   3815: 'Spare_Fault_3815', class No Acknowledgement, trigger "DB302_HMI_Faults_Carrier59_Faults_2" bit 6
   3816: 'Spare_Fault_3816', class No Acknowledgement, trigger "DB302_HMI_Faults_Carrier59_Faults_2" bit 7
   3817: 'Spare_Fault_3817', class No Acknowledgement, trigger "DB302_HMI_Faults_Carrier59_Faults_2" bit 8
   3818: 'Spare_Fault_3818', class No Acknowledgement, trigger "DB302_HMI_Faults_Carrier59_Faults_2" bit 9
   3819: 'Spare_Fault_3819', class No Acknowledgement, trigger "DB302_HMI_Faults_Carrier59_Faults_2" bit 10
   3820: 'Spare_Fault_3820', class No Acknowledgement, trigger "DB302_HMI_Faults_Carrier59_Faults_2" bit 11
   3821: 'Spare_Fault_3821', class No Acknowledgement, trigger "DB302_HMI_Faults_Carrier59_Faults_2" bit 12
   3822: 'Spare_Fault_3822', class No Acknowledgement, trigger "DB302_HMI_Faults_Carrier59_Faults_2" bit 13
   3823: 'Spare_Fault_3823', class No Acknowledgement, trigger "DB302_HMI_Faults_Carrier59_Faults_2" bit 14
   3824: 'Spare_Fault_3824', class No Acknowledgement, trigger "DB302_HMI_Faults_Carrier59_Faults_2" bit 15
   3825: 'Spare_Fault_3825', class No Acknowledgement, trigger "DB302_HMI_Faults_Carrier59_Faults_3" bit 0
   3826: 'Spare_Fault_3826', class No Acknowledgement, trigger "DB302_HMI_Faults_Carrier59_Faults_3" bit 1
   3827: 'Spare_Fault_3827', class No Acknowledgement, trigger "DB302_HMI_Faults_Carrier59_Faults_3" bit 2
   3828: 'Spare_Fault_3828', class No Acknowledgement, trigger "DB302_HMI_Faults_Carrier59_Faults_3" bit 3
   3829: 'Spare_Fault_3829', class No Acknowledgement, trigger "DB302_HMI_Faults_Carrier59_Faults_3" bit 4
   3830: 'Spare_Fault_3830', class No Acknowledgement, trigger "DB302_HMI_Faults_Carrier59_Faults_3" bit 5
   3831: 'Spare_Fault_3831', class No Acknowledgement, trigger "DB302_HMI_Faults_Carrier59_Faults_3" bit 6
   3832: 'Spare_Fault_3832', class No Acknowledgement, trigger "DB302_HMI_Faults_Carrier59_Faults_3" bit 7
   3833: 'Spare_Fault_3833', class No Acknowledgement, trigger "DB302_HMI_Faults_Carrier59_Faults_3" bit 8
   3834: 'Spare_Fault_3834', class No Acknowledgement, trigger "DB302_HMI_Faults_Carrier59_Faults_3" bit 9
   3835: 'Spare_Fault_3835', class No Acknowledgement, trigger "DB302_HMI_Faults_Carrier59_Faults_3" bit 10
   3836: 'Spare_Fault_3836', class No Acknowledgement, trigger "DB302_HMI_Faults_Carrier59_Faults_3" bit 11
   3837: 'Spare_Fault_3837', class No Acknowledgement, trigger "DB302_HMI_Faults_Carrier59_Faults_3" bit 12
   3838: 'Spare_Fault_3838', class No Acknowledgement, trigger "DB302_HMI_Faults_Carrier59_Faults_3" bit 13
   3839: 'Spare_Fault_3839', class No Acknowledgement, trigger "DB302_HMI_Faults_Carrier59_Faults_3" bit 14
   3840: 'Spare_Fault_3840', class No Acknowledgement, trigger "DB302_HMI_Faults_Carrier59_Faults_3" bit 15
   3841: 'Carrier 60 Disconnect Open Power Fault DI11.0', class No Acknowledgement, trigger "DB302_HMI_Faults_Carrier60_Faults_0" bit 0
   3842: 'Carrier 60 Drive Profinet Comm Fault', class No Acknowledgement, trigger "DB302_HMI_Faults_Carrier60_Faults_0" bit 1
   3843: 'Carrier 60 Production Stop Not Reset', class No Acknowledgement, trigger "DB302_HMI_Faults_Carrier60_Faults_0" bit 2
   3844: 'Carrier 60 CB02122 Tripped', class No Acknowledgement, trigger "DB302_HMI_Faults_Carrier60_Faults_0" bit 3
   3845: 'Carrier 60 CB02123 Tripped', class No Acknowledgement, trigger "DB302_HMI_Faults_Carrier60_Faults_0" bit 4
   3846: 'Carrier 60 AUX1 CB Tripped', class No Acknowledgement, trigger "DB302_HMI_Faults_Carrier60_Faults_0" bit 5
   3847: 'Carrier 60 AUX2 CB Tripped', class No Acknowledgement, trigger "DB302_HMI_Faults_Carrier60_Faults_0" bit 6
   3848: 'Carrier 60 PLC Not Communicating', class No Acknowledgement, trigger "DB302_HMI_Faults_Carrier60_Faults_0" bit 7
   3849: 'Carrier 60 Safe Input Card Fault', class No Acknowledgement, trigger "DB302_HMI_Faults_Carrier60_Faults_0" bit 8
   3850: 'Carrier 60 Safe Output Card Fault', class No Acknowledgement, trigger "DB302_HMI_Faults_Carrier60_Faults_0" bit 9
   3851: 'Carrier 60 Standard Input Card Fault', class No Acknowledgement, trigger "DB302_HMI_Faults_Carrier60_Faults_0" bit 10
   3852: 'Carrier 60 Standard Output Card Fault', class No Acknowledgement, trigger "DB302_HMI_Faults_Carrier60_Faults_0" bit 11
   3853: 'Carrier 60 Encoder Position Fault', class No Acknowledgement, trigger "DB302_HMI_Faults_Carrier60_Faults_0" bit 12
   3854: 'Carrier 60 Encoder Internal Error', class No Acknowledgement, trigger "DB302_HMI_Faults_Carrier60_Faults_0" bit 13
   3855: 'Carrier 60 Encoder Comm Fault', class No Acknowledgement, trigger "DB302_HMI_Faults_Carrier60_Faults_0" bit 14
   3856: 'Carrier 60 HMI Comm Fault', class No Acknowledgement, trigger "DB302_HMI_Faults_Carrier60_Faults_0" bit 15
   3857: 'Carrier 60 Crash Detection Fault', class No Acknowledgement, trigger "DB302_HMI_Faults_Carrier60_Faults_1" bit 0
   3858: 'Carrier 60 Carrier Number Invalid', class No Acknowledgement, trigger "DB302_HMI_Faults_Carrier60_Faults_1" bit 1
   3859: 'Carrier 60 Drive: PROFINET configuration error', class No Acknowledgement, trigger "DB302_HMI_Faults_Carrier60_Faults_1" bit 2
   3860: 'Carrier 60 Drive: Error internal communications', class No Acknowledgement, trigger "DB302_HMI_Faults_Carrier60_Faults_1" bit 3
   3861: 'Carrier 60 Drive: Motor overtemperature', class No Acknowledgement, trigger "DB302_HMI_Faults_Carrier60_Faults_1" bit 4
   3862: 'Carrier 60 Drive: Motor overcurrent', class No Acknowledgement, trigger "DB302_HMI_Faults_Carrier60_Faults_1" bit 5
   3863: 'Carrier 60 Drive: Infeed or power unit not ready', class No Acknowledgement, trigger "DB302_HMI_Faults_Carrier60_Faults_1" bit 6
   3864: 'Carrier 60 Drive: Short-circuit/ground fault detected', class No Acknowledgement, trigger "DB302_HMI_Faults_Carrier60_Faults_1" bit 7
   3865: 'Carrier 60 Drive: PROFINET Setpoint timeout', class No Acknowledgement, trigger "DB302_HMI_Faults_Carrier60_Faults_1" bit 8
   3866: 'Carrier 60 Power unit: Overcurrent', class No Acknowledgement, trigger "DB302_HMI_Faults_Carrier60_Faults_1" bit 9
   3867: 'Carrier 60 Power unit: DC link voltage overvoltage', class No Acknowledgement, trigger "DB302_HMI_Faults_Carrier60_Faults_1" bit 10
   3868: 'Carrier 60 Power unit: DC link voltage undervoltage', class No Acknowledgement, trigger "DB302_HMI_Faults_Carrier60_Faults_1" bit 11
   3869: 'Carrier 60 Power unit: Line phase failure in main circuit', class No Acknowledgement, trigger "DB302_HMI_Faults_Carrier60_Faults_1" bit 12
   3870: 'Carrier 60 Power unit: Phase failure motor cable', class No Acknowledgement, trigger "DB302_HMI_Faults_Carrier60_Faults_1" bit 13
   3871: 'Carrier 60 Power unit: Ground fault', class No Acknowledgement, trigger "DB302_HMI_Faults_Carrier60_Faults_1" bit 14
   3872: 'Spare_Fault_3872', class No Acknowledgement, trigger "DB302_HMI_Faults_Carrier60_Faults_1" bit 15
   3873: 'Carrier 60 Motion Off Fault', class No Acknowledgement, trigger "DB302_HMI_Faults_Carrier60_Faults_2" bit 0
   3874: 'Carrier 60 Motion On Fault', class No Acknowledgement, trigger "DB302_HMI_Faults_Carrier60_Faults_2" bit 1
   3875: 'Carrier 60 Spacing Fault', class No Acknowledgement, trigger "DB302_HMI_Faults_Carrier60_Faults_2" bit 2
   3876: 'Carrier 60 Duplicate Carrier Number Fault', class No Acknowledgement, trigger "DB302_HMI_Faults_Carrier60_Faults_2" bit 3
   3877: 'Spare_Fault_3877', class No Acknowledgement, trigger "DB302_HMI_Faults_Carrier60_Faults_2" bit 4
   3878: 'Spare_Fault_3878', class No Acknowledgement, trigger "DB302_HMI_Faults_Carrier60_Faults_2" bit 5
   3879: 'Spare_Fault_3879', class No Acknowledgement, trigger "DB302_HMI_Faults_Carrier60_Faults_2" bit 6
   3880: 'Spare_Fault_3880', class No Acknowledgement, trigger "DB302_HMI_Faults_Carrier60_Faults_2" bit 7
   3881: 'Spare_Fault_3881', class No Acknowledgement, trigger "DB302_HMI_Faults_Carrier60_Faults_2" bit 8
   3882: 'Spare_Fault_3882', class No Acknowledgement, trigger "DB302_HMI_Faults_Carrier60_Faults_2" bit 9
   3883: 'Spare_Fault_3883', class No Acknowledgement, trigger "DB302_HMI_Faults_Carrier60_Faults_2" bit 10
   3884: 'Spare_Fault_3884', class No Acknowledgement, trigger "DB302_HMI_Faults_Carrier60_Faults_2" bit 11
   3885: 'Spare_Fault_3885', class No Acknowledgement, trigger "DB302_HMI_Faults_Carrier60_Faults_2" bit 12
   3886: 'Spare_Fault_3886', class No Acknowledgement, trigger "DB302_HMI_Faults_Carrier60_Faults_2" bit 13
   3887: 'Spare_Fault_3887', class No Acknowledgement, trigger "DB302_HMI_Faults_Carrier60_Faults_2" bit 14
   3888: 'Spare_Fault_3888', class No Acknowledgement, trigger "DB302_HMI_Faults_Carrier60_Faults_2" bit 15
   3889: 'Spare_Fault_3889', class No Acknowledgement, trigger "DB302_HMI_Faults_Carrier60_Faults_3" bit 0
   3890: 'Spare_Fault_3890', class No Acknowledgement, trigger "DB302_HMI_Faults_Carrier60_Faults_3" bit 1
   3891: 'Spare_Fault_3891', class No Acknowledgement, trigger "DB302_HMI_Faults_Carrier60_Faults_3" bit 2
   3892: 'Spare_Fault_3892', class No Acknowledgement, trigger "DB302_HMI_Faults_Carrier60_Faults_3" bit 3
   3893: 'Spare_Fault_3893', class No Acknowledgement, trigger "DB302_HMI_Faults_Carrier60_Faults_3" bit 4
   3894: 'Spare_Fault_3894', class No Acknowledgement, trigger "DB302_HMI_Faults_Carrier60_Faults_3" bit 5
   3895: 'Spare_Fault_3895', class No Acknowledgement, trigger "DB302_HMI_Faults_Carrier60_Faults_3" bit 6
   3896: 'Spare_Fault_3896', class No Acknowledgement, trigger "DB302_HMI_Faults_Carrier60_Faults_3" bit 7
   3897: 'Spare_Fault_3897', class No Acknowledgement, trigger "DB302_HMI_Faults_Carrier60_Faults_3" bit 8
   3898: 'Spare_Fault_3898', class No Acknowledgement, trigger "DB302_HMI_Faults_Carrier60_Faults_3" bit 9
   3899: 'Spare_Fault_3899', class No Acknowledgement, trigger "DB302_HMI_Faults_Carrier60_Faults_3" bit 10
   3900: 'Spare_Fault_3900', class No Acknowledgement, trigger "DB302_HMI_Faults_Carrier60_Faults_3" bit 11
   3901: 'Spare_Fault_3901', class No Acknowledgement, trigger "DB302_HMI_Faults_Carrier60_Faults_3" bit 12
   3902: 'Spare_Fault_3902', class No Acknowledgement, trigger "DB302_HMI_Faults_Carrier60_Faults_3" bit 13
   3903: 'Spare_Fault_3903', class No Acknowledgement, trigger "DB302_HMI_Faults_Carrier60_Faults_3" bit 14
   3904: 'Spare_Fault_3904', class No Acknowledgement, trigger "DB302_HMI_Faults_Carrier60_Faults_3" bit 15
   3905: 'Carrier 61 Disconnect Open Power Fault DI11.0', class No Acknowledgement, trigger "DB302_HMI_Faults_Carrier61_Faults_0" bit 0
   3906: 'Carrier 61 Drive Profinet Comm Fault', class No Acknowledgement, trigger "DB302_HMI_Faults_Carrier61_Faults_0" bit 1
   3907: 'Carrier 61 Production Stop Not Reset', class No Acknowledgement, trigger "DB302_HMI_Faults_Carrier61_Faults_0" bit 2
   3908: 'Carrier 61 CB02122 Tripped', class No Acknowledgement, trigger "DB302_HMI_Faults_Carrier61_Faults_0" bit 3
   3909: 'Carrier 61 CB02123 Tripped', class No Acknowledgement, trigger "DB302_HMI_Faults_Carrier61_Faults_0" bit 4
   3910: 'Carrier 61 AUX1 CB Tripped', class No Acknowledgement, trigger "DB302_HMI_Faults_Carrier61_Faults_0" bit 5
   3911: 'Carrier 61 AUX2 CB Tripped', class No Acknowledgement, trigger "DB302_HMI_Faults_Carrier61_Faults_0" bit 6
   3912: 'Carrier 61 PLC Not Communicating', class No Acknowledgement, trigger "DB302_HMI_Faults_Carrier61_Faults_0" bit 7
   3913: 'Carrier 61 Safe Input Card Fault', class No Acknowledgement, trigger "DB302_HMI_Faults_Carrier61_Faults_0" bit 8
   3914: 'Carrier 61 Safe Output Card Fault', class No Acknowledgement, trigger "DB302_HMI_Faults_Carrier61_Faults_0" bit 9
   3915: 'Carrier 61 Standard Input Card Fault', class No Acknowledgement, trigger "DB302_HMI_Faults_Carrier61_Faults_0" bit 10
   3916: 'Carrier 61 Standard Output Card Fault', class No Acknowledgement, trigger "DB302_HMI_Faults_Carrier61_Faults_0" bit 11
   3917: 'Carrier 61 Encoder Position Fault', class No Acknowledgement, trigger "DB302_HMI_Faults_Carrier61_Faults_0" bit 12
   3918: 'Carrier 61 Encoder Internal Error', class No Acknowledgement, trigger "DB302_HMI_Faults_Carrier61_Faults_0" bit 13
   3919: 'Carrier 61 Encoder Comm Fault', class No Acknowledgement, trigger "DB302_HMI_Faults_Carrier61_Faults_0" bit 14
   3920: 'Carrier 61 HMI Comm Fault', class No Acknowledgement, trigger "DB302_HMI_Faults_Carrier61_Faults_0" bit 15
   3921: 'Carrier 61 Crash Detection Fault', class No Acknowledgement, trigger "DB302_HMI_Faults_Carrier61_Faults_1" bit 0
   3922: 'Carrier 61 Carrier Number Invalid', class No Acknowledgement, trigger "DB302_HMI_Faults_Carrier61_Faults_1" bit 1
   3923: 'Carrier 61 Drive: PROFINET configuration error', class No Acknowledgement, trigger "DB302_HMI_Faults_Carrier61_Faults_1" bit 2
   3924: 'Carrier 61 Drive: Error internal communications', class No Acknowledgement, trigger "DB302_HMI_Faults_Carrier61_Faults_1" bit 3
   3925: 'Carrier 61 Drive: Motor overtemperature', class No Acknowledgement, trigger "DB302_HMI_Faults_Carrier61_Faults_1" bit 4
   3926: 'Carrier 61 Drive: Motor overcurrent', class No Acknowledgement, trigger "DB302_HMI_Faults_Carrier61_Faults_1" bit 5
   3927: 'Carrier 61 Drive: Infeed or power unit not ready', class No Acknowledgement, trigger "DB302_HMI_Faults_Carrier61_Faults_1" bit 6
   3928: 'Carrier 61 Drive: Short-circuit/ground fault detected', class No Acknowledgement, trigger "DB302_HMI_Faults_Carrier61_Faults_1" bit 7
   3929: 'Carrier 61 Drive: PROFINET Setpoint timeout', class No Acknowledgement, trigger "DB302_HMI_Faults_Carrier61_Faults_1" bit 8
   3930: 'Carrier 61 Power unit: Overcurrent', class No Acknowledgement, trigger "DB302_HMI_Faults_Carrier61_Faults_1" bit 9
   3931: 'Carrier 61 Power unit: DC link voltage overvoltage', class No Acknowledgement, trigger "DB302_HMI_Faults_Carrier61_Faults_1" bit 10
   3932: 'Carrier 61 Power unit: DC link voltage undervoltage', class No Acknowledgement, trigger "DB302_HMI_Faults_Carrier61_Faults_1" bit 11
   3933: 'Carrier 61 Power unit: Line phase failure in main circuit', class No Acknowledgement, trigger "DB302_HMI_Faults_Carrier61_Faults_1" bit 12
   3934: 'Carrier 61 Power unit: Phase failure motor cable', class No Acknowledgement, trigger "DB302_HMI_Faults_Carrier61_Faults_1" bit 13
   3935: 'Carrier 61 Power unit: Ground fault', class No Acknowledgement, trigger "DB302_HMI_Faults_Carrier61_Faults_1" bit 14
   3936: 'Spare_Fault_3936', class No Acknowledgement, trigger "DB302_HMI_Faults_Carrier61_Faults_1" bit 15
   3937: 'Carrier 61 Motion Off Fault', class No Acknowledgement, trigger "DB302_HMI_Faults_Carrier61_Faults_2" bit 0
   3938: 'Carrier 61 Motion On Fault', class No Acknowledgement, trigger "DB302_HMI_Faults_Carrier61_Faults_2" bit 1
   3939: 'Carrier 61 Spacing Fault', class No Acknowledgement, trigger "DB302_HMI_Faults_Carrier61_Faults_2" bit 2
   3940: 'Carrier 61 Duplicate Carrier Number Fault', class No Acknowledgement, trigger "DB302_HMI_Faults_Carrier61_Faults_2" bit 3
   3941: 'Spare_Fault_3941', class No Acknowledgement, trigger "DB302_HMI_Faults_Carrier61_Faults_2" bit 4
   3942: 'Spare_Fault_3942', class No Acknowledgement, trigger "DB302_HMI_Faults_Carrier61_Faults_2" bit 5
   3943: 'Spare_Fault_3943', class No Acknowledgement, trigger "DB302_HMI_Faults_Carrier61_Faults_2" bit 6
   3944: 'Spare_Fault_3944', class No Acknowledgement, trigger "DB302_HMI_Faults_Carrier61_Faults_2" bit 7
   3945: 'Spare_Fault_3945', class No Acknowledgement, trigger "DB302_HMI_Faults_Carrier61_Faults_2" bit 8
   3946: 'Spare_Fault_3946', class No Acknowledgement, trigger "DB302_HMI_Faults_Carrier61_Faults_2" bit 9
   3947: 'Spare_Fault_3947', class No Acknowledgement, trigger "DB302_HMI_Faults_Carrier61_Faults_2" bit 10
   3948: 'Spare_Fault_3948', class No Acknowledgement, trigger "DB302_HMI_Faults_Carrier61_Faults_2" bit 11
   3949: 'Spare_Fault_3949', class No Acknowledgement, trigger "DB302_HMI_Faults_Carrier61_Faults_2" bit 12
   3950: 'Spare_Fault_3950', class No Acknowledgement, trigger "DB302_HMI_Faults_Carrier61_Faults_2" bit 13
   3951: 'Spare_Fault_3951', class No Acknowledgement, trigger "DB302_HMI_Faults_Carrier61_Faults_2" bit 14
   3952: 'Spare_Fault_3952', class No Acknowledgement, trigger "DB302_HMI_Faults_Carrier61_Faults_2" bit 15
   3953: 'Spare_Fault_3953', class No Acknowledgement, trigger "DB302_HMI_Faults_Carrier61_Faults_3" bit 0
   3954: 'Spare_Fault_3954', class No Acknowledgement, trigger "DB302_HMI_Faults_Carrier61_Faults_3" bit 1
   3955: 'Spare_Fault_3955', class No Acknowledgement, trigger "DB302_HMI_Faults_Carrier61_Faults_3" bit 2
   3956: 'Spare_Fault_3956', class No Acknowledgement, trigger "DB302_HMI_Faults_Carrier61_Faults_3" bit 3
   3957: 'Spare_Fault_3957', class No Acknowledgement, trigger "DB302_HMI_Faults_Carrier61_Faults_3" bit 4
   3958: 'Spare_Fault_3958', class No Acknowledgement, trigger "DB302_HMI_Faults_Carrier61_Faults_3" bit 5
   3959: 'Spare_Fault_3959', class No Acknowledgement, trigger "DB302_HMI_Faults_Carrier61_Faults_3" bit 6
   3960: 'Spare_Fault_3960', class No Acknowledgement, trigger "DB302_HMI_Faults_Carrier61_Faults_3" bit 7
   3961: 'Spare_Fault_3961', class No Acknowledgement, trigger "DB302_HMI_Faults_Carrier61_Faults_3" bit 8
   3962: 'Spare_Fault_3962', class No Acknowledgement, trigger "DB302_HMI_Faults_Carrier61_Faults_3" bit 9
   3963: 'Spare_Fault_3963', class No Acknowledgement, trigger "DB302_HMI_Faults_Carrier61_Faults_3" bit 10
   3964: 'Spare_Fault_3964', class No Acknowledgement, trigger "DB302_HMI_Faults_Carrier61_Faults_3" bit 11
   3965: 'Spare_Fault_3965', class No Acknowledgement, trigger "DB302_HMI_Faults_Carrier61_Faults_3" bit 12
   3966: 'Spare_Fault_3966', class No Acknowledgement, trigger "DB302_HMI_Faults_Carrier61_Faults_3" bit 13
   3967: 'Spare_Fault_3967', class No Acknowledgement, trigger "DB302_HMI_Faults_Carrier61_Faults_3" bit 14
   3968: 'Spare_Fault_3968', class No Acknowledgement, trigger "DB302_HMI_Faults_Carrier61_Faults_3" bit 15
   3969: 'Carrier 62 Disconnect Open Power Fault DI11.0', class No Acknowledgement, trigger "DB302_HMI_Faults_Carrier62_Faults_0" bit 0
   3970: 'Carrier 62 Drive Profinet Comm Fault', class No Acknowledgement, trigger "DB302_HMI_Faults_Carrier62_Faults_0" bit 1
   3971: 'Carrier 62 Production Stop Not Reset', class No Acknowledgement, trigger "DB302_HMI_Faults_Carrier62_Faults_0" bit 2
   3972: 'Carrier 62 CB02122 Tripped', class No Acknowledgement, trigger "DB302_HMI_Faults_Carrier62_Faults_0" bit 3
   3973: 'Carrier 62 CB02123 Tripped', class No Acknowledgement, trigger "DB302_HMI_Faults_Carrier62_Faults_0" bit 4
   3974: 'Carrier 62 AUX1 CB Tripped', class No Acknowledgement, trigger "DB302_HMI_Faults_Carrier62_Faults_0" bit 5
   3975: 'Carrier 62 AUX2 CB Tripped', class No Acknowledgement, trigger "DB302_HMI_Faults_Carrier62_Faults_0" bit 6
   3976: 'Carrier 62 PLC Not Communicating', class No Acknowledgement, trigger "DB302_HMI_Faults_Carrier62_Faults_0" bit 7
   3977: 'Carrier 62 Safe Input Card Fault', class No Acknowledgement, trigger "DB302_HMI_Faults_Carrier62_Faults_0" bit 8
   3978: 'Carrier 62 Safe Output Card Fault', class No Acknowledgement, trigger "DB302_HMI_Faults_Carrier62_Faults_0" bit 9
   3979: 'Carrier 62 Standard Input Card Fault', class No Acknowledgement, trigger "DB302_HMI_Faults_Carrier62_Faults_0" bit 10
   3980: 'Carrier 62 Standard Output Card Fault', class No Acknowledgement, trigger "DB302_HMI_Faults_Carrier62_Faults_0" bit 11
   3981: 'Carrier 62 Encoder Position Fault', class No Acknowledgement, trigger "DB302_HMI_Faults_Carrier62_Faults_0" bit 12
   3982: 'Carrier 62 Encoder Internal Error', class No Acknowledgement, trigger "DB302_HMI_Faults_Carrier62_Faults_0" bit 13
   3983: 'Carrier 62 Encoder Comm Fault', class No Acknowledgement, trigger "DB302_HMI_Faults_Carrier62_Faults_0" bit 14
   3984: 'Carrier 62 HMI Comm Fault', class No Acknowledgement, trigger "DB302_HMI_Faults_Carrier62_Faults_0" bit 15
   3985: 'Carrier 62 Crash Detection Fault', class No Acknowledgement, trigger "DB302_HMI_Faults_Carrier62_Faults_1" bit 0
   3986: 'Carrier 62 Carrier Number Invalid', class No Acknowledgement, trigger "DB302_HMI_Faults_Carrier62_Faults_1" bit 1
   3987: 'Carrier 62 Drive: PROFINET configuration error', class No Acknowledgement, trigger "DB302_HMI_Faults_Carrier62_Faults_1" bit 2
   3988: 'Carrier 62 Drive: Error internal communications', class No Acknowledgement, trigger "DB302_HMI_Faults_Carrier62_Faults_1" bit 3
   3989: 'Carrier 62 Drive: Motor overtemperature', class No Acknowledgement, trigger "DB302_HMI_Faults_Carrier62_Faults_1" bit 4
   3990: 'Carrier 62 Drive: Motor overcurrent', class No Acknowledgement, trigger "DB302_HMI_Faults_Carrier62_Faults_1" bit 5
   3991: 'Carrier 62 Drive: Infeed or power unit not ready', class No Acknowledgement, trigger "DB302_HMI_Faults_Carrier62_Faults_1" bit 6
   3992: 'Carrier 62 Drive: Short-circuit/ground fault detected', class No Acknowledgement, trigger "DB302_HMI_Faults_Carrier62_Faults_1" bit 7
   3993: 'Carrier 62 Drive: PROFINET Setpoint timeout', class No Acknowledgement, trigger "DB302_HMI_Faults_Carrier62_Faults_1" bit 8
   3994: 'Carrier 62 Power unit: Overcurrent', class No Acknowledgement, trigger "DB302_HMI_Faults_Carrier62_Faults_1" bit 9
   3995: 'Carrier 62 Power unit: DC link voltage overvoltage', class No Acknowledgement, trigger "DB302_HMI_Faults_Carrier62_Faults_1" bit 10
   3996: 'Carrier 62 Power unit: DC link voltage undervoltage', class No Acknowledgement, trigger "DB302_HMI_Faults_Carrier62_Faults_1" bit 11
   3997: 'Carrier 62 Power unit: Line phase failure in main circuit', class No Acknowledgement, trigger "DB302_HMI_Faults_Carrier62_Faults_1" bit 12
   3998: 'Carrier 62 Power unit: Phase failure motor cable', class No Acknowledgement, trigger "DB302_HMI_Faults_Carrier62_Faults_1" bit 13
   3999: 'Carrier 62 Power unit: Ground fault', class No Acknowledgement, trigger "DB302_HMI_Faults_Carrier62_Faults_1" bit 14
   4000: 'Spare_Fault_4000', class No Acknowledgement, trigger "DB302_HMI_Faults_Carrier62_Faults_1" bit 15
   4001: 'Carrier 62 Motion Off Fault', class No Acknowledgement, trigger "DB302_HMI_Faults_Carrier62_Faults_2" bit 0
   4002: 'Carrier 62 Motion On Fault', class No Acknowledgement, trigger "DB302_HMI_Faults_Carrier62_Faults_2" bit 1
   4003: 'Carrier 62 Spacing Fault', class No Acknowledgement, trigger "DB302_HMI_Faults_Carrier62_Faults_2" bit 2
   4004: 'Carrier 62 Duplicate Carrier Number Fault', class No Acknowledgement, trigger "DB302_HMI_Faults_Carrier62_Faults_2" bit 3
   4005: 'Spare_Fault_4005', class No Acknowledgement, trigger "DB302_HMI_Faults_Carrier62_Faults_2" bit 4
   4006: 'Spare_Fault_4006', class No Acknowledgement, trigger "DB302_HMI_Faults_Carrier62_Faults_2" bit 5
   4007: 'Spare_Fault_4007', class No Acknowledgement, trigger "DB302_HMI_Faults_Carrier62_Faults_2" bit 6
   4008: 'Spare_Fault_4008', class No Acknowledgement, trigger "DB302_HMI_Faults_Carrier62_Faults_2" bit 7
   4009: 'Spare_Fault_4009', class No Acknowledgement, trigger "DB302_HMI_Faults_Carrier62_Faults_2" bit 8
   4010: 'Spare_Fault_4010', class No Acknowledgement, trigger "DB302_HMI_Faults_Carrier62_Faults_2" bit 9
   4011: 'Spare_Fault_4011', class No Acknowledgement, trigger "DB302_HMI_Faults_Carrier62_Faults_2" bit 10
   4012: 'Spare_Fault_4012', class No Acknowledgement, trigger "DB302_HMI_Faults_Carrier62_Faults_2" bit 11
   4013: 'Spare_Fault_4013', class No Acknowledgement, trigger "DB302_HMI_Faults_Carrier62_Faults_2" bit 12
   4014: 'Spare_Fault_4014', class No Acknowledgement, trigger "DB302_HMI_Faults_Carrier62_Faults_2" bit 13
   4015: 'Spare_Fault_4015', class No Acknowledgement, trigger "DB302_HMI_Faults_Carrier62_Faults_2" bit 14
   4016: 'Spare_Fault_4016', class No Acknowledgement, trigger "DB302_HMI_Faults_Carrier62_Faults_2" bit 15
   4017: 'Spare_Fault_4017', class No Acknowledgement, trigger "DB302_HMI_Faults_Carrier62_Faults_3" bit 0
   4018: 'Spare_Fault_4018', class No Acknowledgement, trigger "DB302_HMI_Faults_Carrier62_Faults_3" bit 1
   4019: 'Spare_Fault_4019', class No Acknowledgement, trigger "DB302_HMI_Faults_Carrier62_Faults_3" bit 2
   4020: 'Spare_Fault_4020', class No Acknowledgement, trigger "DB302_HMI_Faults_Carrier62_Faults_3" bit 3
   4021: 'Spare_Fault_4021', class No Acknowledgement, trigger "DB302_HMI_Faults_Carrier62_Faults_3" bit 4
   4022: 'Spare_Fault_4022', class No Acknowledgement, trigger "DB302_HMI_Faults_Carrier62_Faults_3" bit 5
   4023: 'Spare_Fault_4023', class No Acknowledgement, trigger "DB302_HMI_Faults_Carrier62_Faults_3" bit 6
   4024: 'Spare_Fault_4024', class No Acknowledgement, trigger "DB302_HMI_Faults_Carrier62_Faults_3" bit 7
   4025: 'Spare_Fault_4025', class No Acknowledgement, trigger "DB302_HMI_Faults_Carrier62_Faults_3" bit 8
   4026: 'Spare_Fault_4026', class No Acknowledgement, trigger "DB302_HMI_Faults_Carrier62_Faults_3" bit 9
   4027: 'Spare_Fault_4027', class No Acknowledgement, trigger "DB302_HMI_Faults_Carrier62_Faults_3" bit 10
   4028: 'Spare_Fault_4028', class No Acknowledgement, trigger "DB302_HMI_Faults_Carrier62_Faults_3" bit 11
   4029: 'Spare_Fault_4029', class No Acknowledgement, trigger "DB302_HMI_Faults_Carrier62_Faults_3" bit 12
   4030: 'Spare_Fault_4030', class No Acknowledgement, trigger "DB302_HMI_Faults_Carrier62_Faults_3" bit 13
   4031: 'Spare_Fault_4031', class No Acknowledgement, trigger "DB302_HMI_Faults_Carrier62_Faults_3" bit 14
   4032: 'Spare_Fault_4032', class No Acknowledgement, trigger "DB302_HMI_Faults_Carrier62_Faults_3" bit 15
   4033: 'Carrier 63 Disconnect Open Power Fault DI11.0', class No Acknowledgement, trigger "DB302_HMI_Faults_Carrier63_Faults_0" bit 0
   4034: 'Carrier 63 Drive Profinet Comm Fault', class No Acknowledgement, trigger "DB302_HMI_Faults_Carrier63_Faults_0" bit 1
   4035: 'Carrier 63 Production Stop Not Reset', class No Acknowledgement, trigger "DB302_HMI_Faults_Carrier63_Faults_0" bit 2
   4036: 'Carrier 63 CB02122 Tripped', class No Acknowledgement, trigger "DB302_HMI_Faults_Carrier63_Faults_0" bit 3
   4037: 'Carrier 63 CB02123 Tripped', class No Acknowledgement, trigger "DB302_HMI_Faults_Carrier63_Faults_0" bit 4
   4038: 'Carrier 63 AUX1 CB Tripped', class No Acknowledgement, trigger "DB302_HMI_Faults_Carrier63_Faults_0" bit 5
   4039: 'Carrier 63 AUX2 CB Tripped', class No Acknowledgement, trigger "DB302_HMI_Faults_Carrier63_Faults_0" bit 6
   4040: 'Carrier 63 PLC Not Communicating', class No Acknowledgement, trigger "DB302_HMI_Faults_Carrier63_Faults_0" bit 7
   4041: 'Carrier 63 Safe Input Card Fault', class No Acknowledgement, trigger "DB302_HMI_Faults_Carrier63_Faults_0" bit 8
   4042: 'Carrier 63 Safe Output Card Fault', class No Acknowledgement, trigger "DB302_HMI_Faults_Carrier63_Faults_0" bit 9
   4043: 'Carrier 63 Standard Input Card Fault', class No Acknowledgement, trigger "DB302_HMI_Faults_Carrier63_Faults_0" bit 10
   4044: 'Carrier 63 Standard Output Card Fault', class No Acknowledgement, trigger "DB302_HMI_Faults_Carrier63_Faults_0" bit 11
   4045: 'Carrier 63 Encoder Position Fault', class No Acknowledgement, trigger "DB302_HMI_Faults_Carrier63_Faults_0" bit 12
   4046: 'Carrier 63 Encoder Internal Error', class No Acknowledgement, trigger "DB302_HMI_Faults_Carrier63_Faults_0" bit 13
   4047: 'Carrier 63 Encoder Comm Fault', class No Acknowledgement, trigger "DB302_HMI_Faults_Carrier63_Faults_0" bit 14
   4048: 'Carrier 63 HMI Comm Fault', class No Acknowledgement, trigger "DB302_HMI_Faults_Carrier63_Faults_0" bit 15
   4049: 'Carrier 63 Crash Detection Fault', class No Acknowledgement, trigger "DB302_HMI_Faults_Carrier63_Faults_1" bit 0
   4050: 'Carrier 63 Carrier Number Invalid', class No Acknowledgement, trigger "DB302_HMI_Faults_Carrier63_Faults_1" bit 1
   4051: 'Carrier 63 Drive: PROFINET configuration error', class No Acknowledgement, trigger "DB302_HMI_Faults_Carrier63_Faults_1" bit 2
   4052: 'Carrier 63 Drive: Error internal communications', class No Acknowledgement, trigger "DB302_HMI_Faults_Carrier63_Faults_1" bit 3
   4053: 'Carrier 63 Drive: Motor overtemperature', class No Acknowledgement, trigger "DB302_HMI_Faults_Carrier63_Faults_1" bit 4
   4054: 'Carrier 63 Drive: Motor overcurrent', class No Acknowledgement, trigger "DB302_HMI_Faults_Carrier63_Faults_1" bit 5
   4055: 'Carrier 63 Drive: Infeed or power unit not ready', class No Acknowledgement, trigger "DB302_HMI_Faults_Carrier63_Faults_1" bit 6
   4056: 'Carrier 63 Drive: Short-circuit/ground fault detected', class No Acknowledgement, trigger "DB302_HMI_Faults_Carrier63_Faults_1" bit 7
   4057: 'Carrier 63 Drive: PROFINET Setpoint timeout', class No Acknowledgement, trigger "DB302_HMI_Faults_Carrier63_Faults_1" bit 8
   4058: 'Carrier 63 Power unit: Overcurrent', class No Acknowledgement, trigger "DB302_HMI_Faults_Carrier63_Faults_1" bit 9
   4059: 'Carrier 63 Power unit: DC link voltage overvoltage', class No Acknowledgement, trigger "DB302_HMI_Faults_Carrier63_Faults_1" bit 10
   4060: 'Carrier 63 Power unit: DC link voltage undervoltage', class No Acknowledgement, trigger "DB302_HMI_Faults_Carrier63_Faults_1" bit 11
   4061: 'Carrier 63 Power unit: Line phase failure in main circuit', class No Acknowledgement, trigger "DB302_HMI_Faults_Carrier63_Faults_1" bit 12
   4062: 'Carrier 63 Power unit: Phase failure motor cable', class No Acknowledgement, trigger "DB302_HMI_Faults_Carrier63_Faults_1" bit 13
   4063: 'Carrier 63 Power unit: Ground fault', class No Acknowledgement, trigger "DB302_HMI_Faults_Carrier63_Faults_1" bit 14
   4064: 'Spare_Fault_4064', class No Acknowledgement, trigger "DB302_HMI_Faults_Carrier63_Faults_1" bit 15
   4065: 'Carrier 63 Motion Off Fault', class No Acknowledgement, trigger "DB302_HMI_Faults_Carrier63_Faults_2" bit 0
   4066: 'Carrier 63 Motion On Fault', class No Acknowledgement, trigger "DB302_HMI_Faults_Carrier63_Faults_2" bit 1
   4067: 'Carrier 63 Spacing Fault', class No Acknowledgement, trigger "DB302_HMI_Faults_Carrier63_Faults_2" bit 2
   4068: 'Carrier 63 Duplicate Carrier Number Fault', class No Acknowledgement, trigger "DB302_HMI_Faults_Carrier63_Faults_2" bit 3
   4069: 'Spare_Fault_4069', class No Acknowledgement, trigger "DB302_HMI_Faults_Carrier63_Faults_2" bit 4
   4070: 'Spare_Fault_4070', class No Acknowledgement, trigger "DB302_HMI_Faults_Carrier63_Faults_2" bit 5
   4071: 'Spare_Fault_4071', class No Acknowledgement, trigger "DB302_HMI_Faults_Carrier63_Faults_2" bit 6
   4072: 'Spare_Fault_4072', class No Acknowledgement, trigger "DB302_HMI_Faults_Carrier63_Faults_2" bit 7
   4073: 'Spare_Fault_4073', class No Acknowledgement, trigger "DB302_HMI_Faults_Carrier63_Faults_2" bit 8
   4074: 'Spare_Fault_4074', class No Acknowledgement, trigger "DB302_HMI_Faults_Carrier63_Faults_2" bit 9
   4075: 'Spare_Fault_4075', class No Acknowledgement, trigger "DB302_HMI_Faults_Carrier63_Faults_2" bit 10
   4076: 'Spare_Fault_4076', class No Acknowledgement, trigger "DB302_HMI_Faults_Carrier63_Faults_2" bit 11
   4077: 'Spare_Fault_4077', class No Acknowledgement, trigger "DB302_HMI_Faults_Carrier63_Faults_2" bit 12
   4078: 'Spare_Fault_4078', class No Acknowledgement, trigger "DB302_HMI_Faults_Carrier63_Faults_2" bit 13
   4079: 'Spare_Fault_4079', class No Acknowledgement, trigger "DB302_HMI_Faults_Carrier63_Faults_2" bit 14
   4080: 'Spare_Fault_4080', class No Acknowledgement, trigger "DB302_HMI_Faults_Carrier63_Faults_2" bit 15
   4081: 'Spare_Fault_4081', class No Acknowledgement, trigger "DB302_HMI_Faults_Carrier63_Faults_3" bit 0
   4082: 'Spare_Fault_4082', class No Acknowledgement, trigger "DB302_HMI_Faults_Carrier63_Faults_3" bit 1
   4083: 'Spare_Fault_4083', class No Acknowledgement, trigger "DB302_HMI_Faults_Carrier63_Faults_3" bit 2
   4084: 'Spare_Fault_4084', class No Acknowledgement, trigger "DB302_HMI_Faults_Carrier63_Faults_3" bit 3
   4085: 'Spare_Fault_4085', class No Acknowledgement, trigger "DB302_HMI_Faults_Carrier63_Faults_3" bit 4
   4086: 'Spare_Fault_4086', class No Acknowledgement, trigger "DB302_HMI_Faults_Carrier63_Faults_3" bit 5
   4087: 'Spare_Fault_4087', class No Acknowledgement, trigger "DB302_HMI_Faults_Carrier63_Faults_3" bit 6
   4088: 'Spare_Fault_4088', class No Acknowledgement, trigger "DB302_HMI_Faults_Carrier63_Faults_3" bit 7
   4089: 'Spare_Fault_4089', class No Acknowledgement, trigger "DB302_HMI_Faults_Carrier63_Faults_3" bit 8
   4090: 'Spare_Fault_4090', class No Acknowledgement, trigger "DB302_HMI_Faults_Carrier63_Faults_3" bit 9
   4091: 'Spare_Fault_4091', class No Acknowledgement, trigger "DB302_HMI_Faults_Carrier63_Faults_3" bit 10
   4092: 'Spare_Fault_4092', class No Acknowledgement, trigger "DB302_HMI_Faults_Carrier63_Faults_3" bit 11
   4093: 'Spare_Fault_4093', class No Acknowledgement, trigger "DB302_HMI_Faults_Carrier63_Faults_3" bit 12
   4094: 'Spare_Fault_4094', class No Acknowledgement, trigger "DB302_HMI_Faults_Carrier63_Faults_3" bit 13
   4095: 'Spare_Fault_4095', class No Acknowledgement, trigger "DB302_HMI_Faults_Carrier63_Faults_3" bit 14
   4096: 'Spare_Fault_4096', class No Acknowledgement, trigger "DB302_HMI_Faults_Carrier63_Faults_3" bit 15
   4097: 'Carrier 64 Disconnect Open Power Fault DI11.0', class No Acknowledgement, trigger "DB302_HMI_Faults_Carrier64_Faults_0" bit 0
   4098: 'Carrier 64 Drive Profinet Comm Fault', class No Acknowledgement, trigger "DB302_HMI_Faults_Carrier64_Faults_0" bit 1
   4099: 'Carrier 64 Production Stop Not Reset', class No Acknowledgement, trigger "DB302_HMI_Faults_Carrier64_Faults_0" bit 2
   4100: 'Carrier 64 CB02122 Tripped', class No Acknowledgement, trigger "DB302_HMI_Faults_Carrier64_Faults_0" bit 3
   4101: 'Carrier 64 CB02123 Tripped', class No Acknowledgement, trigger "DB302_HMI_Faults_Carrier64_Faults_0" bit 4
   4102: 'Carrier 64 AUX1 CB Tripped', class No Acknowledgement, trigger "DB302_HMI_Faults_Carrier64_Faults_0" bit 5
   4103: 'Carrier 64 AUX2 CB Tripped', class No Acknowledgement, trigger "DB302_HMI_Faults_Carrier64_Faults_0" bit 6
   4104: 'Carrier 64 PLC Not Communicating', class No Acknowledgement, trigger "DB302_HMI_Faults_Carrier64_Faults_0" bit 7
   4105: 'Carrier 64 Safe Input Card Fault', class No Acknowledgement, trigger "DB302_HMI_Faults_Carrier64_Faults_0" bit 8
   4106: 'Carrier 64 Safe Output Card Fault', class No Acknowledgement, trigger "DB302_HMI_Faults_Carrier64_Faults_0" bit 9
   4107: 'Carrier 64 Standard Input Card Fault', class No Acknowledgement, trigger "DB302_HMI_Faults_Carrier64_Faults_0" bit 10
   4108: 'Carrier 64 Standard Output Card Fault', class No Acknowledgement, trigger "DB302_HMI_Faults_Carrier64_Faults_0" bit 11
   4109: 'Carrier 64 Encoder Position Fault', class No Acknowledgement, trigger "DB302_HMI_Faults_Carrier64_Faults_0" bit 12
   4110: 'Carrier 64 Encoder Internal Error', class No Acknowledgement, trigger "DB302_HMI_Faults_Carrier64_Faults_0" bit 13
   4111: 'Carrier 64 Encoder Comm Fault', class No Acknowledgement, trigger "DB302_HMI_Faults_Carrier64_Faults_0" bit 14
   4112: 'Carrier 64 HMI Comm Fault', class No Acknowledgement, trigger "DB302_HMI_Faults_Carrier64_Faults_0" bit 15
   4113: 'Carrier 64 Crash Detection Fault', class No Acknowledgement, trigger "DB302_HMI_Faults_Carrier64_Faults_1" bit 0
   4114: 'Carrier 64 Carrier Number Invalid', class No Acknowledgement, trigger "DB302_HMI_Faults_Carrier64_Faults_1" bit 1
   4115: 'Carrier 64 Drive: PROFINET configuration error', class No Acknowledgement, trigger "DB302_HMI_Faults_Carrier64_Faults_1" bit 2
   4116: 'Carrier 64 Drive: Error internal communications', class No Acknowledgement, trigger "DB302_HMI_Faults_Carrier64_Faults_1" bit 3
   4117: 'Carrier 64 Drive: Motor overtemperature', class No Acknowledgement, trigger "DB302_HMI_Faults_Carrier64_Faults_1" bit 4
   4118: 'Carrier 64 Drive: Motor overcurrent', class No Acknowledgement, trigger "DB302_HMI_Faults_Carrier64_Faults_1" bit 5
   4119: 'Carrier 64 Drive: Infeed or power unit not ready', class No Acknowledgement, trigger "DB302_HMI_Faults_Carrier64_Faults_1" bit 6
   4120: 'Carrier 64 Drive: Short-circuit/ground fault detected', class No Acknowledgement, trigger "DB302_HMI_Faults_Carrier64_Faults_1" bit 7
   4121: 'Carrier 64 Drive: PROFINET Setpoint timeout', class No Acknowledgement, trigger "DB302_HMI_Faults_Carrier64_Faults_1" bit 8
   4122: 'Carrier 64 Power unit: Overcurrent', class No Acknowledgement, trigger "DB302_HMI_Faults_Carrier64_Faults_1" bit 9
   4123: 'Carrier 64 Power unit: DC link voltage overvoltage', class No Acknowledgement, trigger "DB302_HMI_Faults_Carrier64_Faults_1" bit 10
   4124: 'Carrier 64 Power unit: DC link voltage undervoltage', class No Acknowledgement, trigger "DB302_HMI_Faults_Carrier64_Faults_1" bit 11
   4125: 'Carrier 64 Power unit: Line phase failure in main circuit', class No Acknowledgement, trigger "DB302_HMI_Faults_Carrier64_Faults_1" bit 12
   4126: 'Carrier 64 Power unit: Phase failure motor cable', class No Acknowledgement, trigger "DB302_HMI_Faults_Carrier64_Faults_1" bit 13
   4127: 'Carrier 64 Power unit: Ground fault', class No Acknowledgement, trigger "DB302_HMI_Faults_Carrier64_Faults_1" bit 14
   4128: 'Spare_Fault_4128', class No Acknowledgement, trigger "DB302_HMI_Faults_Carrier64_Faults_1" bit 15
   4129: 'Carrier 64 Motion Off Fault', class No Acknowledgement, trigger "DB302_HMI_Faults_Carrier64_Faults_2" bit 0
   4130: 'Carrier 64 Motion On Fault', class No Acknowledgement, trigger "DB302_HMI_Faults_Carrier64_Faults_2" bit 1
   4131: 'Carrier 64 Spacing Fault', class No Acknowledgement, trigger "DB302_HMI_Faults_Carrier64_Faults_2" bit 2
   4132: 'Carrier 64 Duplicate Carrier Number Fault', class No Acknowledgement, trigger "DB302_HMI_Faults_Carrier64_Faults_2" bit 3
   4133: 'Spare_Fault_4133', class No Acknowledgement, trigger "DB302_HMI_Faults_Carrier64_Faults_2" bit 4
   4134: 'Spare_Fault_4134', class No Acknowledgement, trigger "DB302_HMI_Faults_Carrier64_Faults_2" bit 5
   4135: 'Spare_Fault_4135', class No Acknowledgement, trigger "DB302_HMI_Faults_Carrier64_Faults_2" bit 6
   4136: 'Spare_Fault_4136', class No Acknowledgement, trigger "DB302_HMI_Faults_Carrier64_Faults_2" bit 7
   4137: 'Spare_Fault_4137', class No Acknowledgement, trigger "DB302_HMI_Faults_Carrier64_Faults_2" bit 8
   4138: 'Spare_Fault_4138', class No Acknowledgement, trigger "DB302_HMI_Faults_Carrier64_Faults_2" bit 9
   4139: 'Spare_Fault_4139', class No Acknowledgement, trigger "DB302_HMI_Faults_Carrier64_Faults_2" bit 10
   4140: 'Spare_Fault_4140', class No Acknowledgement, trigger "DB302_HMI_Faults_Carrier64_Faults_2" bit 11
   4141: 'Spare_Fault_4141', class No Acknowledgement, trigger "DB302_HMI_Faults_Carrier64_Faults_2" bit 12
   4142: 'Spare_Fault_4142', class No Acknowledgement, trigger "DB302_HMI_Faults_Carrier64_Faults_2" bit 13
   4143: 'Spare_Fault_4143', class No Acknowledgement, trigger "DB302_HMI_Faults_Carrier64_Faults_2" bit 14
   4144: 'Spare_Fault_4144', class No Acknowledgement, trigger "DB302_HMI_Faults_Carrier64_Faults_2" bit 15
   4145: 'Spare_Fault_4145', class No Acknowledgement, trigger "DB302_HMI_Faults_Carrier64_Faults_3" bit 0
   4146: 'Spare_Fault_4146', class No Acknowledgement, trigger "DB302_HMI_Faults_Carrier64_Faults_3" bit 1
   4147: 'Spare_Fault_4147', class No Acknowledgement, trigger "DB302_HMI_Faults_Carrier64_Faults_3" bit 2
   4148: 'Spare_Fault_4148', class No Acknowledgement, trigger "DB302_HMI_Faults_Carrier64_Faults_3" bit 3
   4149: 'Spare_Fault_4149', class No Acknowledgement, trigger "DB302_HMI_Faults_Carrier64_Faults_3" bit 4
   4150: 'Spare_Fault_4150', class No Acknowledgement, trigger "DB302_HMI_Faults_Carrier64_Faults_3" bit 5
   4151: 'Spare_Fault_4151', class No Acknowledgement, trigger "DB302_HMI_Faults_Carrier64_Faults_3" bit 6
   4152: 'Spare_Fault_4152', class No Acknowledgement, trigger "DB302_HMI_Faults_Carrier64_Faults_3" bit 7
   4153: 'Spare_Fault_4153', class No Acknowledgement, trigger "DB302_HMI_Faults_Carrier64_Faults_3" bit 8
   4154: 'Spare_Fault_4154', class No Acknowledgement, trigger "DB302_HMI_Faults_Carrier64_Faults_3" bit 9
   4155: 'Spare_Fault_4155', class No Acknowledgement, trigger "DB302_HMI_Faults_Carrier64_Faults_3" bit 10
   4156: 'Spare_Fault_4156', class No Acknowledgement, trigger "DB302_HMI_Faults_Carrier64_Faults_3" bit 11
   4157: 'Spare_Fault_4157', class No Acknowledgement, trigger "DB302_HMI_Faults_Carrier64_Faults_3" bit 12
   4158: 'Spare_Fault_4158', class No Acknowledgement, trigger "DB302_HMI_Faults_Carrier64_Faults_3" bit 13
   4159: 'Spare_Fault_4159', class No Acknowledgement, trigger "DB302_HMI_Faults_Carrier64_Faults_3" bit 14
   4160: 'Spare_Fault_4160', class No Acknowledgement, trigger "DB302_HMI_Faults_Carrier64_Faults_3" bit 15
   4161: 'Carrier 65 Disconnect Open Power Fault DI11.0', class No Acknowledgement, trigger "DB302_HMI_Faults_Carrier65_Faults_0" bit 0
   4162: 'Carrier 65 Drive Profinet Comm Fault', class No Acknowledgement, trigger "DB302_HMI_Faults_Carrier65_Faults_0" bit 1
   4163: 'Carrier 65 Production Stop Not Reset', class No Acknowledgement, trigger "DB302_HMI_Faults_Carrier65_Faults_0" bit 2
   4164: 'Carrier 65 CB02122 Tripped', class No Acknowledgement, trigger "DB302_HMI_Faults_Carrier65_Faults_0" bit 3
   4165: 'Carrier 65 CB02123 Tripped', class No Acknowledgement, trigger "DB302_HMI_Faults_Carrier65_Faults_0" bit 4
   4166: 'Carrier 65 AUX1 CB Tripped', class No Acknowledgement, trigger "DB302_HMI_Faults_Carrier65_Faults_0" bit 5
   4167: 'Carrier 65 AUX2 CB Tripped', class No Acknowledgement, trigger "DB302_HMI_Faults_Carrier65_Faults_0" bit 6
   4168: 'Carrier 65 PLC Not Communicating', class No Acknowledgement, trigger "DB302_HMI_Faults_Carrier65_Faults_0" bit 7
   4169: 'Carrier 65 Safe Input Card Fault', class No Acknowledgement, trigger "DB302_HMI_Faults_Carrier65_Faults_0" bit 8
   4170: 'Carrier 65 Safe Output Card Fault', class No Acknowledgement, trigger "DB302_HMI_Faults_Carrier65_Faults_0" bit 9
   4171: 'Carrier 65 Standard Input Card Fault', class No Acknowledgement, trigger "DB302_HMI_Faults_Carrier65_Faults_0" bit 10
   4172: 'Carrier 65 Standard Output Card Fault', class No Acknowledgement, trigger "DB302_HMI_Faults_Carrier65_Faults_0" bit 11
   4173: 'Carrier 65 Encoder Position Fault', class No Acknowledgement, trigger "DB302_HMI_Faults_Carrier65_Faults_0" bit 12
   4174: 'Carrier 65 Encoder Internal Error', class No Acknowledgement, trigger "DB302_HMI_Faults_Carrier65_Faults_0" bit 13
   4175: 'Carrier 65 Encoder Comm Fault', class No Acknowledgement, trigger "DB302_HMI_Faults_Carrier65_Faults_0" bit 14
   4176: 'Carrier 65 HMI Comm Fault', class No Acknowledgement, trigger "DB302_HMI_Faults_Carrier65_Faults_0" bit 15
   4177: 'Carrier 65 Crash Detection Fault', class No Acknowledgement, trigger "DB302_HMI_Faults_Carrier65_Faults_1" bit 0
   4178: 'Carrier 65 Carrier Number Invalid', class No Acknowledgement, trigger "DB302_HMI_Faults_Carrier65_Faults_1" bit 1
   4179: 'Carrier 65 Drive: PROFINET configuration error', class No Acknowledgement, trigger "DB302_HMI_Faults_Carrier65_Faults_1" bit 2
   4180: 'Carrier 65 Drive: Error internal communications', class No Acknowledgement, trigger "DB302_HMI_Faults_Carrier65_Faults_1" bit 3
   4181: 'Carrier 65 Drive: Motor overtemperature', class No Acknowledgement, trigger "DB302_HMI_Faults_Carrier65_Faults_1" bit 4
   4182: 'Carrier 65 Drive: Motor overcurrent', class No Acknowledgement, trigger "DB302_HMI_Faults_Carrier65_Faults_1" bit 5
   4183: 'Carrier 65 Drive: Infeed or power unit not ready', class No Acknowledgement, trigger "DB302_HMI_Faults_Carrier65_Faults_1" bit 6
   4184: 'Carrier 65 Drive: Short-circuit/ground fault detected', class No Acknowledgement, trigger "DB302_HMI_Faults_Carrier65_Faults_1" bit 7
   4185: 'Carrier 65 Drive: PROFINET Setpoint timeout', class No Acknowledgement, trigger "DB302_HMI_Faults_Carrier65_Faults_1" bit 8
   4186: 'Carrier 65 Power unit: Overcurrent', class No Acknowledgement, trigger "DB302_HMI_Faults_Carrier65_Faults_1" bit 9
   4187: 'Carrier 65 Power unit: DC link voltage overvoltage', class No Acknowledgement, trigger "DB302_HMI_Faults_Carrier65_Faults_1" bit 10
   4188: 'Carrier 65 Power unit: DC link voltage undervoltage', class No Acknowledgement, trigger "DB302_HMI_Faults_Carrier65_Faults_1" bit 11
   4189: 'Carrier 65 Power unit: Line phase failure in main circuit', class No Acknowledgement, trigger "DB302_HMI_Faults_Carrier65_Faults_1" bit 12
   4190: 'Carrier 65 Power unit: Phase failure motor cable', class No Acknowledgement, trigger "DB302_HMI_Faults_Carrier65_Faults_1" bit 13
   4191: 'Carrier 65 Power unit: Ground fault', class No Acknowledgement, trigger "DB302_HMI_Faults_Carrier65_Faults_1" bit 14
   4192: 'Spare_Fault_4192', class No Acknowledgement, trigger "DB302_HMI_Faults_Carrier65_Faults_1" bit 15
   4193: 'Carrier 65 Motion Off Fault', class No Acknowledgement, trigger "DB302_HMI_Faults_Carrier65_Faults_2" bit 0
   4194: 'Carrier 65 Motion On Fault', class No Acknowledgement, trigger "DB302_HMI_Faults_Carrier65_Faults_2" bit 1
   4195: 'Carrier 65 Spacing Fault', class No Acknowledgement, trigger "DB302_HMI_Faults_Carrier65_Faults_2" bit 2
   4196: 'Carrier 65 Duplicate Carrier Number Fault', class No Acknowledgement, trigger "DB302_HMI_Faults_Carrier65_Faults_2" bit 3
   4197: 'Spare_Fault_4197', class No Acknowledgement, trigger "DB302_HMI_Faults_Carrier65_Faults_2" bit 4
   4198: 'Spare_Fault_4198', class No Acknowledgement, trigger "DB302_HMI_Faults_Carrier65_Faults_2" bit 5
   4199: 'Spare_Fault_4199', class No Acknowledgement, trigger "DB302_HMI_Faults_Carrier65_Faults_2" bit 6
   4200: 'Spare_Fault_4200', class No Acknowledgement, trigger "DB302_HMI_Faults_Carrier65_Faults_2" bit 7
   4201: 'Spare_Fault_4201', class No Acknowledgement, trigger "DB302_HMI_Faults_Carrier65_Faults_2" bit 8
   4202: 'Spare_Fault_4202', class No Acknowledgement, trigger "DB302_HMI_Faults_Carrier65_Faults_2" bit 9
   4203: 'Spare_Fault_4203', class No Acknowledgement, trigger "DB302_HMI_Faults_Carrier65_Faults_2" bit 10
   4204: 'Spare_Fault_4204', class No Acknowledgement, trigger "DB302_HMI_Faults_Carrier65_Faults_2" bit 11
   4205: 'Spare_Fault_4205', class No Acknowledgement, trigger "DB302_HMI_Faults_Carrier65_Faults_2" bit 12
   4206: 'Spare_Fault_4206', class No Acknowledgement, trigger "DB302_HMI_Faults_Carrier65_Faults_2" bit 13
   4207: 'Spare_Fault_4207', class No Acknowledgement, trigger "DB302_HMI_Faults_Carrier65_Faults_2" bit 14
   4208: 'Spare_Fault_4208', class No Acknowledgement, trigger "DB302_HMI_Faults_Carrier65_Faults_2" bit 15
   4209: 'Spare_Fault_4209', class No Acknowledgement, trigger "DB302_HMI_Faults_Carrier65_Faults_3" bit 0
   4210: 'Spare_Fault_4210', class No Acknowledgement, trigger "DB302_HMI_Faults_Carrier65_Faults_3" bit 1
   4211: 'Spare_Fault_4211', class No Acknowledgement, trigger "DB302_HMI_Faults_Carrier65_Faults_3" bit 2
   4212: 'Spare_Fault_4212', class No Acknowledgement, trigger "DB302_HMI_Faults_Carrier65_Faults_3" bit 3
   4213: 'Spare_Fault_4213', class No Acknowledgement, trigger "DB302_HMI_Faults_Carrier65_Faults_3" bit 4
   4214: 'Spare_Fault_4214', class No Acknowledgement, trigger "DB302_HMI_Faults_Carrier65_Faults_3" bit 5
   4215: 'Spare_Fault_4215', class No Acknowledgement, trigger "DB302_HMI_Faults_Carrier65_Faults_3" bit 6
   4216: 'Spare_Fault_4216', class No Acknowledgement, trigger "DB302_HMI_Faults_Carrier65_Faults_3" bit 7
   4217: 'Spare_Fault_4217', class No Acknowledgement, trigger "DB302_HMI_Faults_Carrier65_Faults_3" bit 8
   4218: 'Spare_Fault_4218', class No Acknowledgement, trigger "DB302_HMI_Faults_Carrier65_Faults_3" bit 9
   4219: 'Spare_Fault_4219', class No Acknowledgement, trigger "DB302_HMI_Faults_Carrier65_Faults_3" bit 10
   4220: 'Spare_Fault_4220', class No Acknowledgement, trigger "DB302_HMI_Faults_Carrier65_Faults_3" bit 11
   4221: 'Spare_Fault_4221', class No Acknowledgement, trigger "DB302_HMI_Faults_Carrier65_Faults_3" bit 12
   4222: 'Spare_Fault_4222', class No Acknowledgement, trigger "DB302_HMI_Faults_Carrier65_Faults_3" bit 13
   4223: 'Spare_Fault_4223', class No Acknowledgement, trigger "DB302_HMI_Faults_Carrier65_Faults_3" bit 14
   4224: 'Spare_Fault_4224', class No Acknowledgement, trigger "DB302_HMI_Faults_Carrier65_Faults_3" bit 15
   4225: 'Carrier 66 Disconnect Open Power Fault DI11.0', class No Acknowledgement, trigger "DB302_HMI_Faults_Carrier66_Faults_0" bit 0
   4226: 'Carrier 66 Drive Profinet Comm Fault', class No Acknowledgement, trigger "DB302_HMI_Faults_Carrier66_Faults_0" bit 1
   4227: 'Carrier 66 Production Stop Not Reset', class No Acknowledgement, trigger "DB302_HMI_Faults_Carrier66_Faults_0" bit 2
   4228: 'Carrier 66 CB02122 Tripped', class No Acknowledgement, trigger "DB302_HMI_Faults_Carrier66_Faults_0" bit 3
   4229: 'Carrier 66 CB02123 Tripped', class No Acknowledgement, trigger "DB302_HMI_Faults_Carrier66_Faults_0" bit 4
   4230: 'Carrier 66 AUX1 CB Tripped', class No Acknowledgement, trigger "DB302_HMI_Faults_Carrier66_Faults_0" bit 5
   4231: 'Carrier 66 AUX2 CB Tripped', class No Acknowledgement, trigger "DB302_HMI_Faults_Carrier66_Faults_0" bit 6
   4232: 'Carrier 66 PLC Not Communicating', class No Acknowledgement, trigger "DB302_HMI_Faults_Carrier66_Faults_0" bit 7
   4233: 'Carrier 66 Safe Input Card Fault', class No Acknowledgement, trigger "DB302_HMI_Faults_Carrier66_Faults_0" bit 8
   4234: 'Carrier 66 Safe Output Card Fault', class No Acknowledgement, trigger "DB302_HMI_Faults_Carrier66_Faults_0" bit 9
   4235: 'Carrier 66 Standard Input Card Fault', class No Acknowledgement, trigger "DB302_HMI_Faults_Carrier66_Faults_0" bit 10
   4236: 'Carrier 66 Standard Output Card Fault', class No Acknowledgement, trigger "DB302_HMI_Faults_Carrier66_Faults_0" bit 11
   4237: 'Carrier 66 Encoder Position Fault', class No Acknowledgement, trigger "DB302_HMI_Faults_Carrier66_Faults_0" bit 12
